(* Logix 5000 project; controller _GigaDiscovery vendor 1 type 14 code 244 rev 35.11; software revision 35.03; part 6 of 23 *)
(* tags used below, declared in another part *)
   Encoder_Pulses : DINT;
   Pignone : DINT;
   Pylon_Axe_Position_360_SUB : REAL;
   Ralla : DINT;
   RallaPignone : REAL;
   Riduttore : REAL;
   Timer : TIMER[50];
   Clock : DINT;   // Base tempi 10 milli sec
   Clock_1_Hz : BOOL;   // SL Clock 1 Hz 0.5 sec OFF 0.5 sec ON
   Clock_4_Hz : BOOL;   // SL Clock 4 Hz 0.125 sec OFF 0.125 sec ON
   Emergency_Brake_manual_Perm : BOOL;
   Emergency_Brake_SL : ALIAS FOR K300_OCC:6:O.6;   // _S31207D
   Gates_Open_Permissive : Permissive;
   Gondola_Axe : Axe;
   HMI_Lamp_Test : BOOL;
   HMI_Monitor_Bars_Time : DINT;
   I_EStop_Pb_OCC1 : UDT_DCI_STOP_TEST;   // +OCC E-stop -S30301F
   I_EStop_Pb_OCC2 : UDT_DCI_STOP_TEST;   // +OCC2 E-Stop -S28502F
   I_Gate_2_Opened : BOOL;   // Gate 2 RFID Sensor Closed -B24601J
   I_Gate_3_Opened : BOOL;   // Gate 3 RFID Sensor Closed -B24701J
   I_Gate_ENTER_G01_Closed : UDT_DCM;   // GATE ENTER (G01) -B25204I
   I_Gate_EXIT_G05_Closed : UDT_DCM;   // GATE EXIT (G05) -B25304I
   I_OCC1_Stop_Cycle_PB : BOOL;   // Stop Cycle -S30308F
   I_OCC2_ACONFIRM : BOOL;   // OCC2 Allow Main CONFIRM -S28602F
   I_OCC2_Stop_Cycle_PB : BOOL;   // Stop Cycle -S28606F
   I_OCC_Emergency_Brake : BOOL;   // I OCC Emergency Brake -S31207D
   I_OCC_Operator_Enable_Key : BOOL;   // OCC Console Enabled -S30305F
   I_Zero_Set_Sensor : BOOL;   // Zero Set Sensor -B11201A
   Impulsi_per_360_gradi : DINT;
   Impulsi_per_grado : REAL;
   K_Speed_Factor : REAL;
   Mem_RESTRAINTS_closed_Correctly : BOOL;
   MODE : BOOL;   // MODE 0 = AUTO 1 = MANUAL -S30801F
   No_Emergencies_CL0 : BOOL;
   No_Emergencies_CL1 : BOOL;
   No_Sfty : Std_to_Sfty;
   O_Close_Gate2 : BOOL;   // Gate 2 Exit Close = Mag ON
   O_Close_Gate3 : BOOL;   // Gate 3 Entrance Close = Mag ON
   O_OCC_EStop_SL : ALIAS FOR K300_OCC:5:O.7;   // -S30301F EMERGENCY
   O_Start_Signal_2 : ALIAS FOR K300_OCC:5:O.2;   // -S30401F RIDE START
   Pb_Platform_Stop : BOOL;   // Platform Stop Command -S30608F
   Platform_Close_Cycle : Sequencer;
   Platform_Close_Permissive_OK : BOOL;
   Platform_Closed_Aux : DINT;
   Platform_Open_Cycle : Sequencer;
   Platform_Open_Permissive : Permissive;
   Platform_Open_Permissive_Ok : BOOL;
   Platform_Opened_Aux : DINT;
   PltaformClosed_CycleComplete : BOOL;   // Piattaforme chiuse e ciclo completato
   PltaformOpeneded_CycleComplete : BOOL;   // Rilevazione Piattaforme aperte con ciclo Completato
   Pylon_Axe : Axe;
   Pylon_Filtered_Speed : REAL;
   Pylon_Filtered_Speed_ABS : REAL;
   Pylon_Stop_Phase : BOOL;
   Reset_Status_SL_Request : BOOL;
   RESTRAINTS_Closed : BOOL;   // All RESTRAINTS Closed
   RESTRAINTS_Open_Postion : BOOL[64];
   RESTRAINTS_Sector : LapBars_Sector[9];
   Start_Platform_AutoCycle_Pylon : BOOL;
   Start_Stop_Cycle : Sequencer;
   Timers : TIMER[32];
   To_Sfty : Std_to_Sfty;
(* Input, continued *)

ROUTINE _04_RESTRAINTS   (* ladder *)
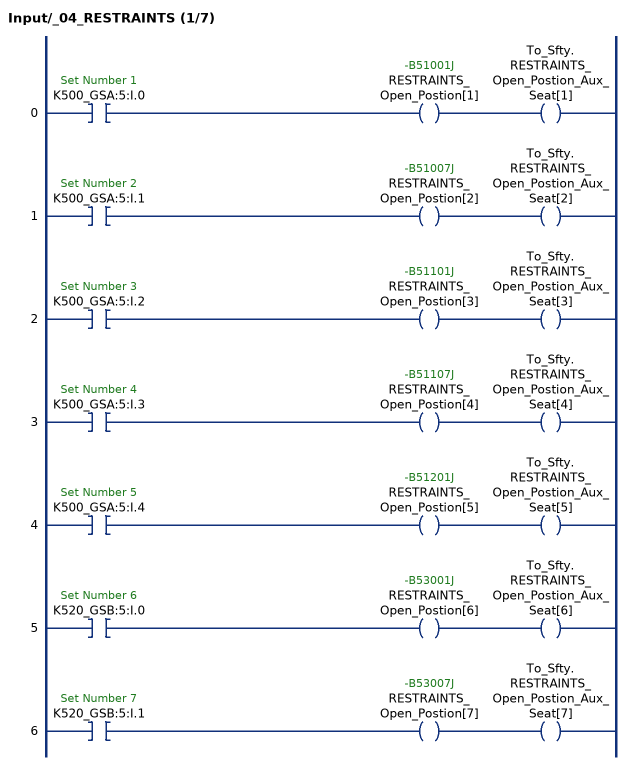
   0: XIC(K500_GSA:5:I.0)OTE(RESTRAINTS_Open_Postion[1])OTE(To_Sfty.RESTRAINTS_Open_Postion_Aux_Seat[1]);
   1: XIC(K500_GSA:5:I.1)OTE(RESTRAINTS_Open_Postion[2])OTE(To_Sfty.RESTRAINTS_Open_Postion_Aux_Seat[2]);
   2: XIC(K500_GSA:5:I.2)OTE(RESTRAINTS_Open_Postion[3])OTE(To_Sfty.RESTRAINTS_Open_Postion_Aux_Seat[3]);
   3: XIC(K500_GSA:5:I.3)OTE(RESTRAINTS_Open_Postion[4])OTE(To_Sfty.RESTRAINTS_Open_Postion_Aux_Seat[4]);
   4: XIC(K500_GSA:5:I.4)OTE(RESTRAINTS_Open_Postion[5])OTE(To_Sfty.RESTRAINTS_Open_Postion_Aux_Seat[5]);
   5: XIC(K520_GSB:5:I.0)OTE(RESTRAINTS_Open_Postion[6])OTE(To_Sfty.RESTRAINTS_Open_Postion_Aux_Seat[6]);
   6: XIC(K520_GSB:5:I.1)OTE(RESTRAINTS_Open_Postion[7])OTE(To_Sfty.RESTRAINTS_Open_Postion_Aux_Seat[7]);
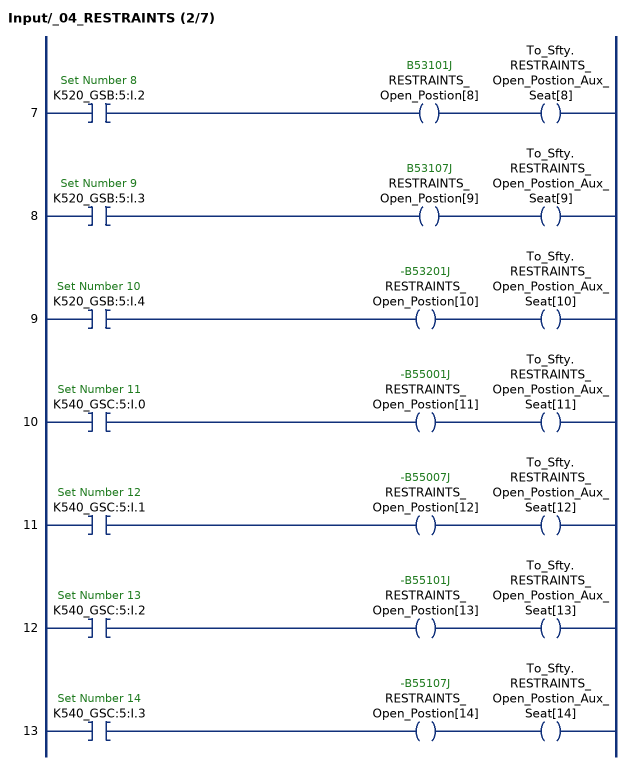
   7: XIC(K520_GSB:5:I.2)OTE(RESTRAINTS_Open_Postion[8])OTE(To_Sfty.RESTRAINTS_Open_Postion_Aux_Seat[8]);
   8: XIC(K520_GSB:5:I.3)OTE(RESTRAINTS_Open_Postion[9])OTE(To_Sfty.RESTRAINTS_Open_Postion_Aux_Seat[9]);
   9: XIC(K520_GSB:5:I.4)OTE(RESTRAINTS_Open_Postion[10])OTE(To_Sfty.RESTRAINTS_Open_Postion_Aux_Seat[10]);
   10: XIC(K540_GSC:5:I.0)OTE(RESTRAINTS_Open_Postion[11])OTE(To_Sfty.RESTRAINTS_Open_Postion_Aux_Seat[11]);
   11: XIC(K540_GSC:5:I.1)OTE(RESTRAINTS_Open_Postion[12])OTE(To_Sfty.RESTRAINTS_Open_Postion_Aux_Seat[12]);
   12: XIC(K540_GSC:5:I.2)OTE(RESTRAINTS_Open_Postion[13])OTE(To_Sfty.RESTRAINTS_Open_Postion_Aux_Seat[13]);
   13: XIC(K540_GSC:5:I.3)OTE(RESTRAINTS_Open_Postion[14])OTE(To_Sfty.RESTRAINTS_Open_Postion_Aux_Seat[14]);
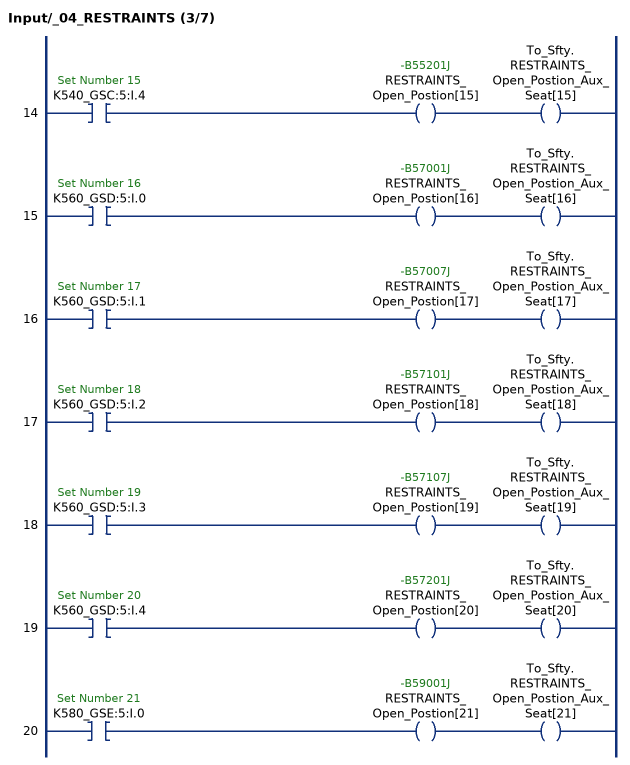
   14: XIC(K540_GSC:5:I.4)OTE(RESTRAINTS_Open_Postion[15])OTE(To_Sfty.RESTRAINTS_Open_Postion_Aux_Seat[15]);
   15: XIC(K560_GSD:5:I.0)OTE(RESTRAINTS_Open_Postion[16])OTE(To_Sfty.RESTRAINTS_Open_Postion_Aux_Seat[16]);
   16: XIC(K560_GSD:5:I.1)OTE(RESTRAINTS_Open_Postion[17])OTE(To_Sfty.RESTRAINTS_Open_Postion_Aux_Seat[17]);
   17: XIC(K560_GSD:5:I.2)OTE(RESTRAINTS_Open_Postion[18])OTE(To_Sfty.RESTRAINTS_Open_Postion_Aux_Seat[18]);
   18: XIC(K560_GSD:5:I.3)OTE(RESTRAINTS_Open_Postion[19])OTE(To_Sfty.RESTRAINTS_Open_Postion_Aux_Seat[19]);
   19: XIC(K560_GSD:5:I.4)OTE(RESTRAINTS_Open_Postion[20])OTE(To_Sfty.RESTRAINTS_Open_Postion_Aux_Seat[20]);
   20: XIC(K580_GSE:5:I.0)OTE(RESTRAINTS_Open_Postion[21])OTE(To_Sfty.RESTRAINTS_Open_Postion_Aux_Seat[21]);
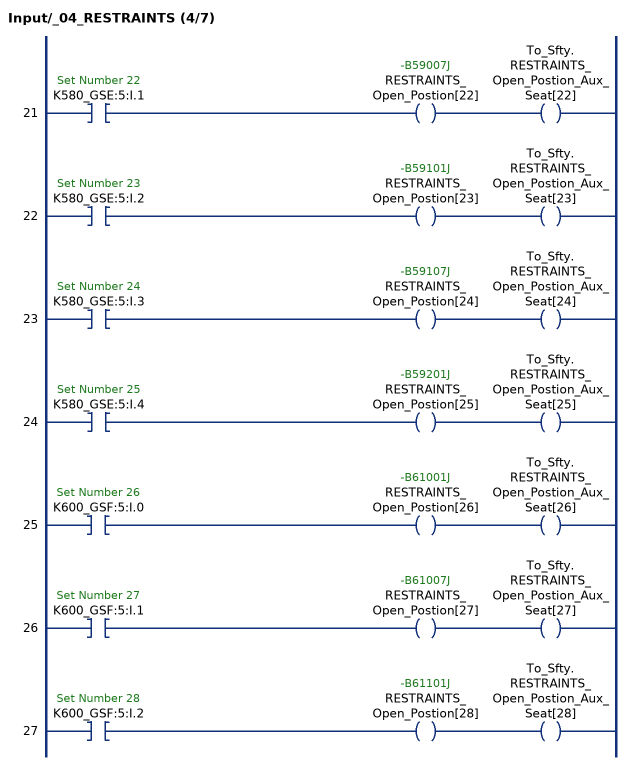
   21: XIC(K580_GSE:5:I.1)OTE(RESTRAINTS_Open_Postion[22])OTE(To_Sfty.RESTRAINTS_Open_Postion_Aux_Seat[22]);
   22: XIC(K580_GSE:5:I.2)OTE(RESTRAINTS_Open_Postion[23])OTE(To_Sfty.RESTRAINTS_Open_Postion_Aux_Seat[23]);
   23: XIC(K580_GSE:5:I.3)OTE(RESTRAINTS_Open_Postion[24])OTE(To_Sfty.RESTRAINTS_Open_Postion_Aux_Seat[24]);
   24: XIC(K580_GSE:5:I.4)OTE(RESTRAINTS_Open_Postion[25])OTE(To_Sfty.RESTRAINTS_Open_Postion_Aux_Seat[25]);
   25: XIC(K600_GSF:5:I.0)OTE(RESTRAINTS_Open_Postion[26])OTE(To_Sfty.RESTRAINTS_Open_Postion_Aux_Seat[26]);
   26: XIC(K600_GSF:5:I.1)OTE(RESTRAINTS_Open_Postion[27])OTE(To_Sfty.RESTRAINTS_Open_Postion_Aux_Seat[27]);
   27: XIC(K600_GSF:5:I.2)OTE(RESTRAINTS_Open_Postion[28])OTE(To_Sfty.RESTRAINTS_Open_Postion_Aux_Seat[28]);
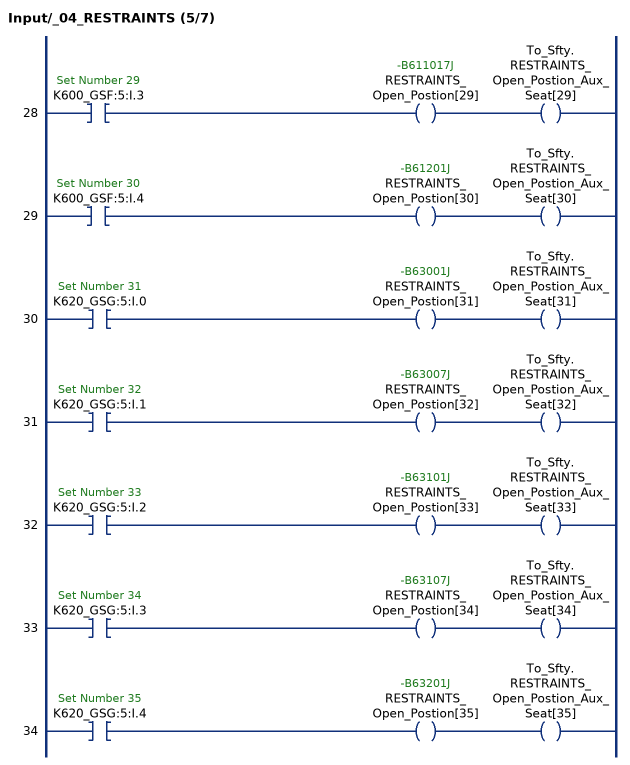
   28: XIC(K600_GSF:5:I.3)OTE(RESTRAINTS_Open_Postion[29])OTE(To_Sfty.RESTRAINTS_Open_Postion_Aux_Seat[29]);
   29: XIC(K600_GSF:5:I.4)OTE(RESTRAINTS_Open_Postion[30])OTE(To_Sfty.RESTRAINTS_Open_Postion_Aux_Seat[30]);
   30: XIC(K620_GSG:5:I.0)OTE(RESTRAINTS_Open_Postion[31])OTE(To_Sfty.RESTRAINTS_Open_Postion_Aux_Seat[31]);
   31: XIC(K620_GSG:5:I.1)OTE(RESTRAINTS_Open_Postion[32])OTE(To_Sfty.RESTRAINTS_Open_Postion_Aux_Seat[32]);
   32: XIC(K620_GSG:5:I.2)OTE(RESTRAINTS_Open_Postion[33])OTE(To_Sfty.RESTRAINTS_Open_Postion_Aux_Seat[33]);
   33: XIC(K620_GSG:5:I.3)OTE(RESTRAINTS_Open_Postion[34])OTE(To_Sfty.RESTRAINTS_Open_Postion_Aux_Seat[34]);
   34: XIC(K620_GSG:5:I.4)OTE(RESTRAINTS_Open_Postion[35])OTE(To_Sfty.RESTRAINTS_Open_Postion_Aux_Seat[35]);
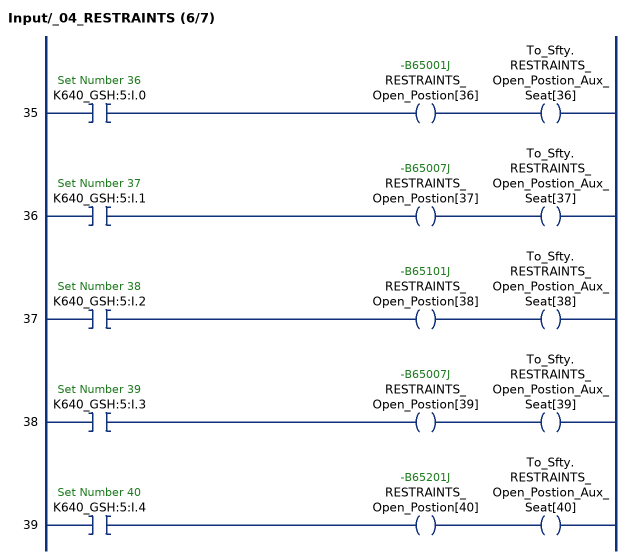
   35: XIC(K640_GSH:5:I.0)OTE(RESTRAINTS_Open_Postion[36])OTE(To_Sfty.RESTRAINTS_Open_Postion_Aux_Seat[36]);
   36: XIC(K640_GSH:5:I.1)OTE(RESTRAINTS_Open_Postion[37])OTE(To_Sfty.RESTRAINTS_Open_Postion_Aux_Seat[37]);
   37: XIC(K640_GSH:5:I.2)OTE(RESTRAINTS_Open_Postion[38])OTE(To_Sfty.RESTRAINTS_Open_Postion_Aux_Seat[38]);
   38: XIC(K640_GSH:5:I.3)OTE(RESTRAINTS_Open_Postion[39])OTE(To_Sfty.RESTRAINTS_Open_Postion_Aux_Seat[39]);
   39: XIC(K640_GSH:5:I.4)OTE(RESTRAINTS_Open_Postion[40])OTE(To_Sfty.RESTRAINTS_Open_Postion_Aux_Seat[40]);
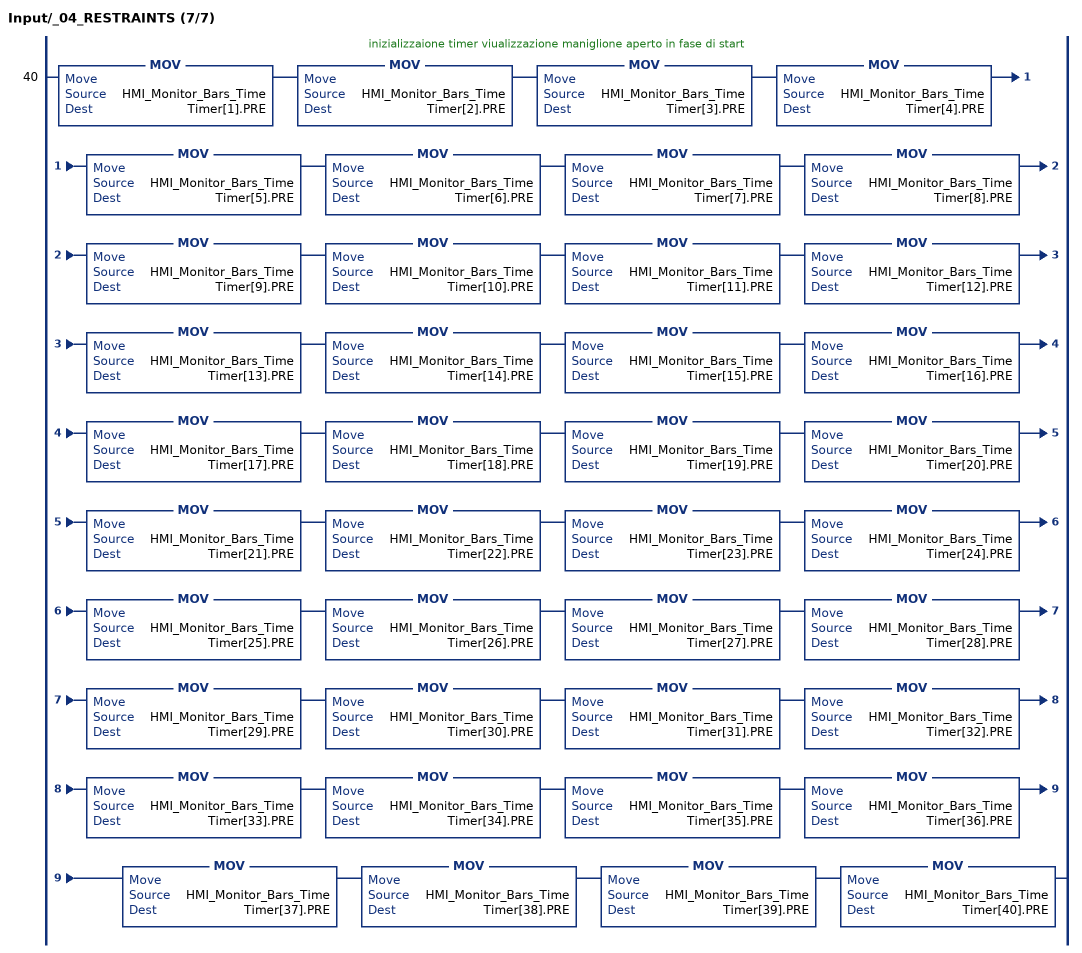
   // inizializzaione timer viualizzazione maniglione aperto in fase di start
   40: MOV(HMI_Monitor_Bars_Time,Timer[1].PRE)MOV(HMI_Monitor_Bars_Time,Timer[2].PRE)MOV(HMI_Monitor_Bars_Time,Timer[3].PRE)MOV(HMI_Monitor_Bars_Time,Timer[4].PRE)MOV(HMI_Monitor_Bars_Time,Timer[5].PRE)MOV(HMI_Monitor_Bars_Time,Timer[6].PRE)MOV(HMI_Monitor_Bars_Time,Timer[7].PRE)MOV(HMI_Monitor_Bars_Time,Timer[8].PRE)MOV(HMI_Monitor_Bars_Time,Timer[9].PRE)MOV(HMI_Monitor_Bars_Time,Timer[10].PRE)MOV(HMI_Monitor_Bars_Time,Timer[11].PRE)MOV(HMI_Monitor_Bars_Time,Timer[12].PRE)MOV(HMI_Monitor_Bars_Time,Timer[13].PRE)MOV(HMI_Monitor_Bars_Time,Timer[14].PRE)MOV(HMI_Monitor_Bars_Time,Timer[15].PRE)MOV(HMI_Monitor_Bars_Time,Timer[16].PRE)MOV(HMI_Monitor_Bars_Time,Timer[17].PRE)MOV(HMI_Monitor_Bars_Time,Timer[18].PRE)MOV(HMI_Monitor_Bars_Time,Timer[19].PRE)MOV(HMI_Monitor_Bars_Time,Timer[20].PRE)MOV(HMI_Monitor_Bars_Time,Timer[21].PRE)MOV(HMI_Monitor_Bars_Time,Timer[22].PRE)MOV(HMI_Monitor_Bars_Time,Timer[23].PRE)MOV(HMI_Monitor_Bars_Time,Timer[24].PRE)MOV(HMI_Monitor_Bars_Time,Timer[25].PRE)MOV(HMI_Monitor_Bars_Time,Timer[26].PRE)MOV(HMI_Monitor_Bars_Time,Timer[27].PRE)MOV(HMI_Monitor_Bars_Time,Timer[28].PRE)MOV(HMI_Monitor_Bars_Time,Timer[29].PRE)MOV(HMI_Monitor_Bars_Time,Timer[30].PRE)MOV(HMI_Monitor_Bars_Time,Timer[31].PRE)MOV(HMI_Monitor_Bars_Time,Timer[32].PRE)MOV(HMI_Monitor_Bars_Time,Timer[33].PRE)MOV(HMI_Monitor_Bars_Time,Timer[34].PRE)MOV(HMI_Monitor_Bars_Time,Timer[35].PRE)MOV(HMI_Monitor_Bars_Time,Timer[36].PRE)MOV(HMI_Monitor_Bars_Time,Timer[37].PRE)MOV(HMI_Monitor_Bars_Time,Timer[38].PRE)MOV(HMI_Monitor_Bars_Time,Timer[39].PRE)MOV(HMI_Monitor_Bars_Time,Timer[40].PRE);
END_ROUTINE

ROUTINE _05_Platform   (* ladder *)
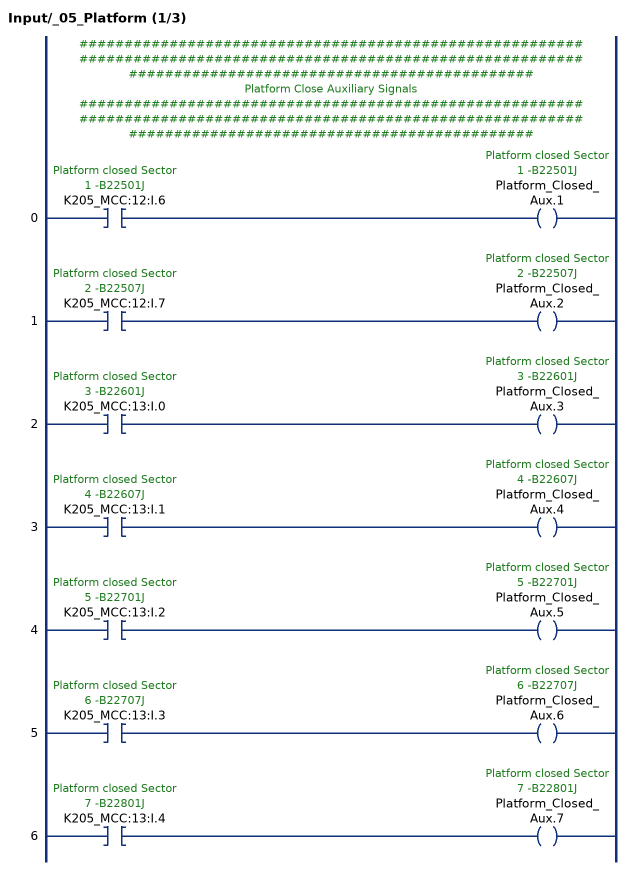
   // #############################################################################################################################################################
   // Platform Close Auxiliary Signals
   // #############################################################################################################################################################
   0: XIC(K205_MCC:12:I.6)OTE(Platform_Closed_Aux.1);
   1: XIC(K205_MCC:12:I.7)OTE(Platform_Closed_Aux.2);
   2: XIC(K205_MCC:13:I.0)OTE(Platform_Closed_Aux.3);
   3: XIC(K205_MCC:13:I.1)OTE(Platform_Closed_Aux.4);
   4: XIC(K205_MCC:13:I.2)OTE(Platform_Closed_Aux.5);
   5: XIC(K205_MCC:13:I.3)OTE(Platform_Closed_Aux.6);
   6: XIC(K205_MCC:13:I.4)OTE(Platform_Closed_Aux.7);
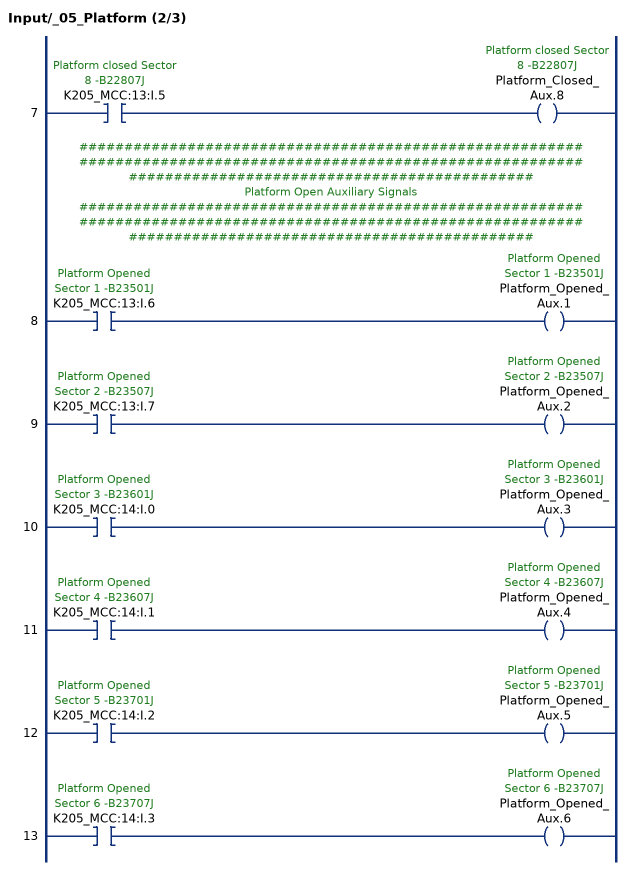
   7: XIC(K205_MCC:13:I.5)OTE(Platform_Closed_Aux.8);
   // #############################################################################################################################################################
   // Platform Open Auxiliary Signals
   // #############################################################################################################################################################
   8: XIC(K205_MCC:13:I.6)OTE(Platform_Opened_Aux.1);
   9: XIC(K205_MCC:13:I.7)OTE(Platform_Opened_Aux.2);
   10: XIC(K205_MCC:14:I.0)OTE(Platform_Opened_Aux.3);
   11: XIC(K205_MCC:14:I.1)OTE(Platform_Opened_Aux.4);
   12: XIC(K205_MCC:14:I.2)OTE(Platform_Opened_Aux.5);
   13: XIC(K205_MCC:14:I.3)OTE(Platform_Opened_Aux.6);
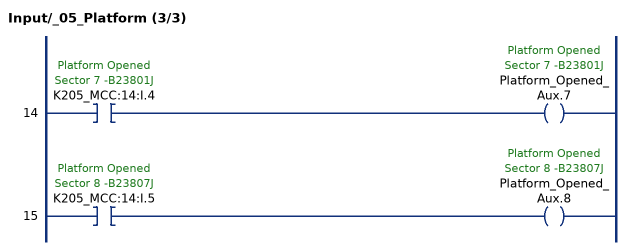
   14: XIC(K205_MCC:14:I.4)OTE(Platform_Opened_Aux.7);
   15: XIC(K205_MCC:14:I.5)OTE(Platform_Opened_Aux.8);
END_ROUTINE

ROUTINE _06_Pylon   (* ladder *)
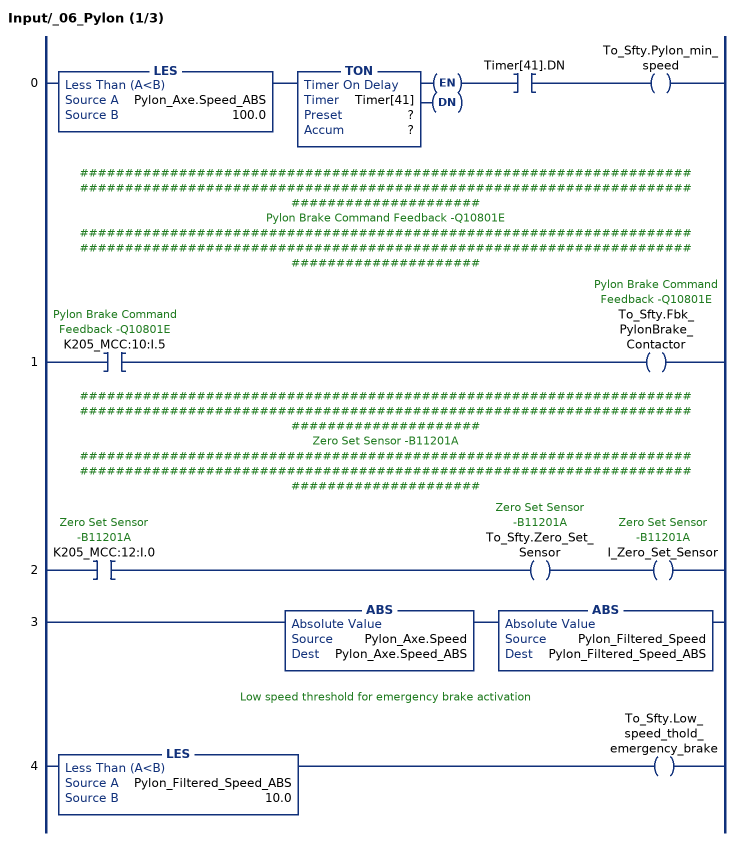
   0: LES(Pylon_Axe.Speed_ABS,100.0)TON(Timer[41],?,?)XIC(Timer[41].DN)OTE(To_Sfty.Pylon_min_speed);
   // #############################################################################################################################################################
   // Pylon Brake Command Feedback -Q10801E
   // #############################################################################################################################################################
   1: XIC(K205_MCC:10:I.5)OTE(To_Sfty.Fbk_PylonBrake_Contactor);
   // #############################################################################################################################################################
   // Zero Set Sensor -B11201A
   // #############################################################################################################################################################
   2: XIC(K205_MCC:12:I.0)OTE(To_Sfty.Zero_Set_Sensor)OTE(I_Zero_Set_Sensor);
   3: ABS(Pylon_Axe.Speed,Pylon_Axe.Speed_ABS)ABS(Pylon_Filtered_Speed,Pylon_Filtered_Speed_ABS);
   // Low speed threshold for emergency brake activation
   4: LES(Pylon_Filtered_Speed_ABS,10.0)OTE(To_Sfty.Low_speed_thold_emergency_brake);
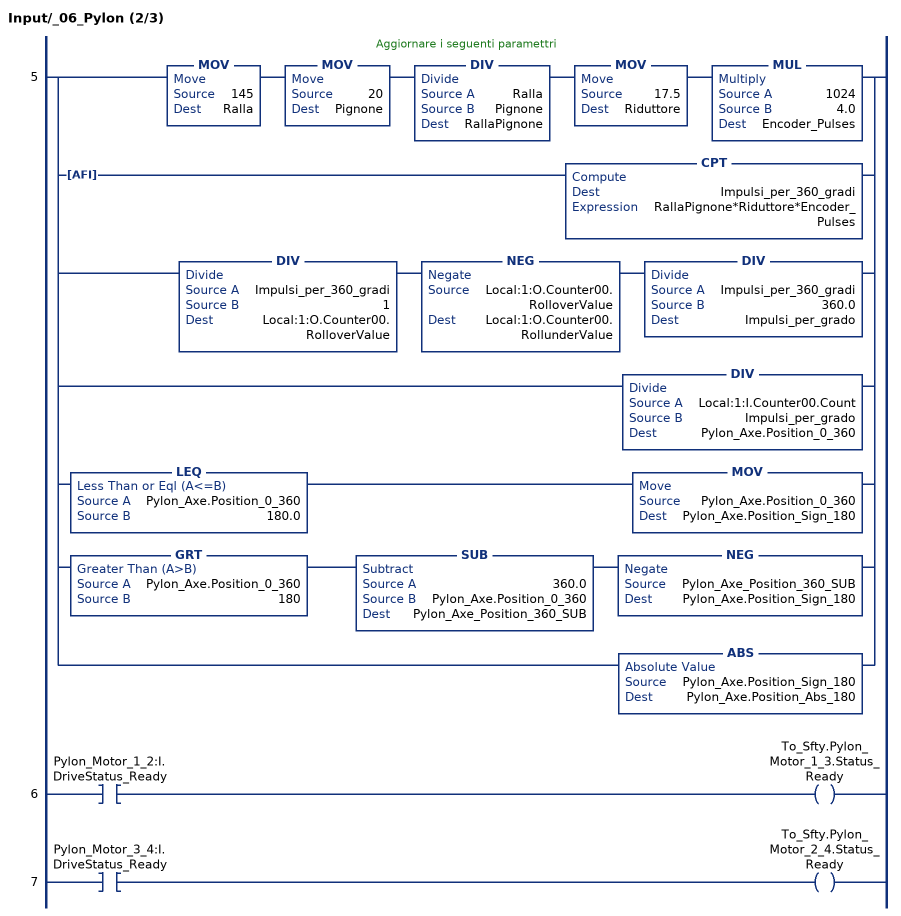
   // Aggiornare i seguenti paramettri
   5: [MOV(145,Ralla) MOV(20,Pignone) DIV(Ralla,Pignone,RallaPignone) MOV(17.5,Riduttore) MUL(1024,4.0,Encoder_Pulses) ,AFI() CPT(Impulsi_per_360_gradi,RallaPignone*Riduttore*Encoder_Pulses) ,DIV(Impulsi_per_360_gradi,1,Local:1:O.Counter00.RolloverValue) NEG(Local:1:O.Counter00.RolloverValue,Local:1:O.Counter00.RollunderValue) DIV(Impulsi_per_360_gradi,360.0,Impulsi_per_grado) ,DIV(Local:1:I.Counter00.Count,Impulsi_per_grado,Pylon_Axe.Position_0_360) ,LEQ(Pylon_Axe.Position_0_360,180.0) MOV(Pylon_Axe.Position_0_360,Pylon_Axe.Position_Sign_180) ,GRT(Pylon_Axe.Position_0_360,180) SUB(360.0,Pylon_Axe.Position_0_360,Pylon_Axe_Position_360_SUB) NEG(Pylon_Axe_Position_360_SUB,Pylon_Axe.Position_Sign_180) ,ABS(Pylon_Axe.Position_Sign_180,Pylon_Axe.Position_Abs_180) ];
   6: XIC(Pylon_Motor_1_2:I.DriveStatus_Ready)OTE(To_Sfty.Pylon_Motor_1_3.Status_Ready);
   7: XIC(Pylon_Motor_3_4:I.DriveStatus_Ready)OTE(To_Sfty.Pylon_Motor_2_4.Status_Ready);
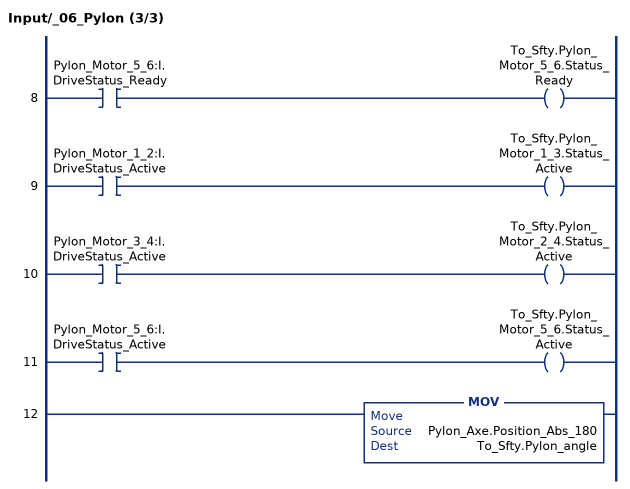
   8: XIC(Pylon_Motor_5_6:I.DriveStatus_Ready)OTE(To_Sfty.Pylon_Motor_5_6.Status_Ready);
   9: XIC(Pylon_Motor_1_2:I.DriveStatus_Active)OTE(To_Sfty.Pylon_Motor_1_3.Status_Active);
   10: XIC(Pylon_Motor_3_4:I.DriveStatus_Active)OTE(To_Sfty.Pylon_Motor_2_4.Status_Active);
   11: XIC(Pylon_Motor_5_6:I.DriveStatus_Active)OTE(To_Sfty.Pylon_Motor_5_6.Status_Active);
   12: MOV(Pylon_Axe.Position_Abs_180,To_Sfty.Pylon_angle);
END_ROUTINE

ROUTINE _07_Gondola   (* ladder *)
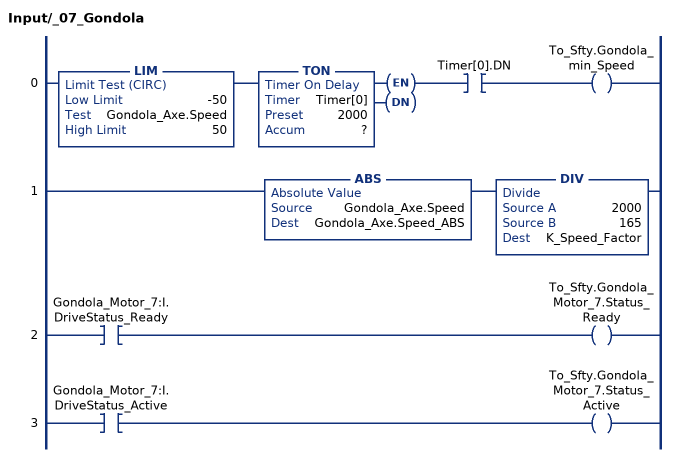
   0: LIM(-50,Gondola_Axe.Speed,50)TON(Timer[0],?,?)XIC(Timer[0].DN)OTE(To_Sfty.Gondola_min_Speed);
   1: ABS(Gondola_Axe.Speed,Gondola_Axe.Speed_ABS)DIV(2000,165,K_Speed_Factor);
   2: XIC(Gondola_Motor_7:I.DriveStatus_Ready)OTE(To_Sfty.Gondola_Motor_7.Status_Ready);
   3: XIC(Gondola_Motor_7:I.DriveStatus_Active)OTE(To_Sfty.Gondola_Motor_7.Status_Active);
END_ROUTINE

ROUTINE Main   (* ladder *)
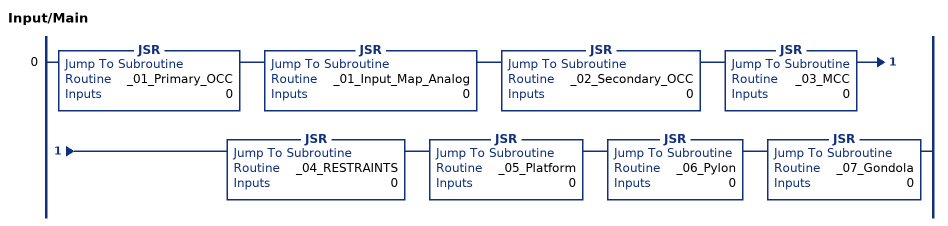
   0: JSR(_01_Primary_OCC,0)JSR(_01_Input_Map_Analog,0)JSR(_02_Secondary_OCC,0)JSR(_03_MCC,0)JSR(_04_RESTRAINTS,0)JSR(_05_Platform,0)JSR(_06_Pylon,0)JSR(_07_Gondola,0);
END_ROUTINE
END_PROGRAM

PROGRAM Main10ms   (* main routine Main *)

ROUTINE Main   (* ladder *)
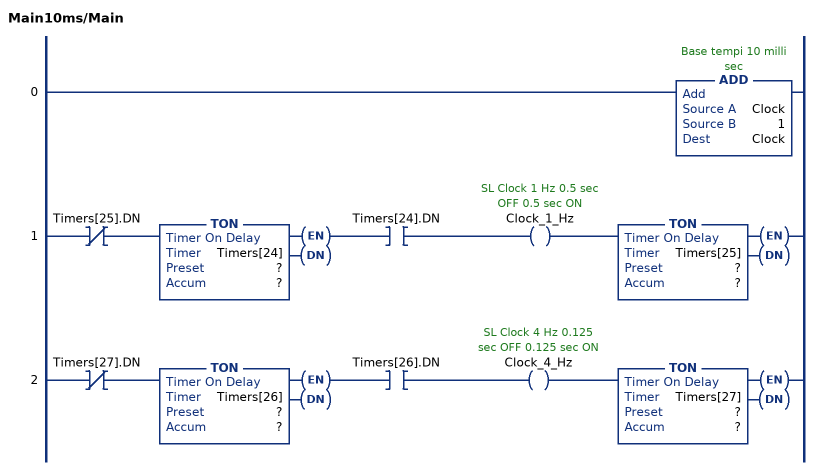
   0: ADD(Clock,1,Clock);
   1: XIO(Timers[25].DN)TON(Timers[24],?,?)XIC(Timers[24].DN)OTE(Clock_1_Hz)TON(Timers[25],?,?);
   2: XIO(Timers[27].DN)TON(Timers[26],?,?)XIC(Timers[26].DN)OTE(Clock_4_Hz)TON(Timers[27],?,?);
END_ROUTINE
END_PROGRAM

PROGRAM Output   (* main routine Main *)
VAR
   EntryGate : Sfq_Lamp := (Input := 1, LampCoil := 1);
   ExitGate : Sfq_Lamp := (Input := 1, LampCoil := 1);
   I_OCC1_Stop_Cycle_PB_memory : BOOL;
   I_OCC2_Stop_Cycle_PB_memory : BOOL;
   O_Alarm_Noise : BOOL;
   O_Alarm_Signal : BOOL;
   O_Allow_Operator : BOOL;
   O_ExitGate_Signal : BOOL := 1;
   O_Lapbars_Open : ALIAS FOR K300_OCC:5:O.4;
   O_Platform_Close_Signal : ALIAS FOR K300_OCC:5:O.6;   // -S30605F PLATFORM CLOSING
   O_Platform_Open_Signal : ALIAS FOR K300_OCC:5:O.5;   // -S30601F PLATFORM OPENING
   O_Start_Signal : ALIAS FOR K300_OCC:5:O.1;   // -S30403F RIDE START
   O_Stop_Signal : ALIAS FOR K300_OCC:5:O.0;   // -S30308F RIDE STOP
   Os : DINT;
   Out_FGEN_01 : FUNCTION_GENERATOR := (XY1Size := 2, Out := -90.0);
   Out_FGEN_06 : FUNCTION_GENERATOR := (XY1Size := 2);
   Out_FGEN_07 : FUNCTION_GENERATOR := (In := -1.0, XY1Size := 2);
   Out_FGEN_09 : FUNCTION_GENERATOR := (XY1Size := 2);
   Out_FGEN_10 : FUNCTION_GENERATOR := (In := 100.0, XY1Size := 2, Out := 10000.0);
   Output_Scalaggi : Scale_2_P[16] := ([0].Input[1] := 100.0, [0].Output[0] := -90.0, [0].Output[1] := 90.0, [1].Input[0] := -100.0, [1].Input[1] := 100.0, [1].Output[0] := -10000.0, [1].Output[1] := 10000.0, [2].Input[1] := 100.0, [2].Output[1] := 10000.0, [3].Input[0] := -100.0, [3].Input[1] := 100.0, [3].Output[0] := -10000.0, [3].Output[1] := 10000.0, [4].Input[1] := 31218.0, [4].Output[1] := 10.0, [5].Input[1] := 31218.0, [5].Output[1] := 10.0, [6].Input[1] := 31218.0, [6].Output[1] := 10.0, [7].Input[1] := 31218.0, [7].Output[1] := 10.0, [8].Input[1] := 31218.0, [8].Output[1] := 10.0, [9].Input[1] := 31218.0, [9].Output[1] := 10.0, [11].Input[0] := -1.0, [11].Input[1] := 1.0, [11].Output[1] := 10000.0, [12].Input[0] := -1.0, [12].Input[1] := 1.0, [12].Output[0] := -10000.0, [12].Output[1] := 10000.0);
   RAD_01 : FBD_MATH_ADVANCED := (Source := -90.0, Dest := -1.5707964);
   SFQ_disable : BOOL;
   SFQ_Mask : DINT := -269484034;
   SFQ_Mask2 : DINT;
   SFQ_MASK_OK : DINT := -1;
   SFQBit : BOOL;
   SIN_01 : FBD_MATH_ADVANCED := (Source := -1.5707964, Dest := -1.0);
   Start_Permissive_MakCompare : DINT := -1048577;
   TempSFQ : DINT;
END_VAR

ROUTINE _01_Primary_OCC   (* ladder *)
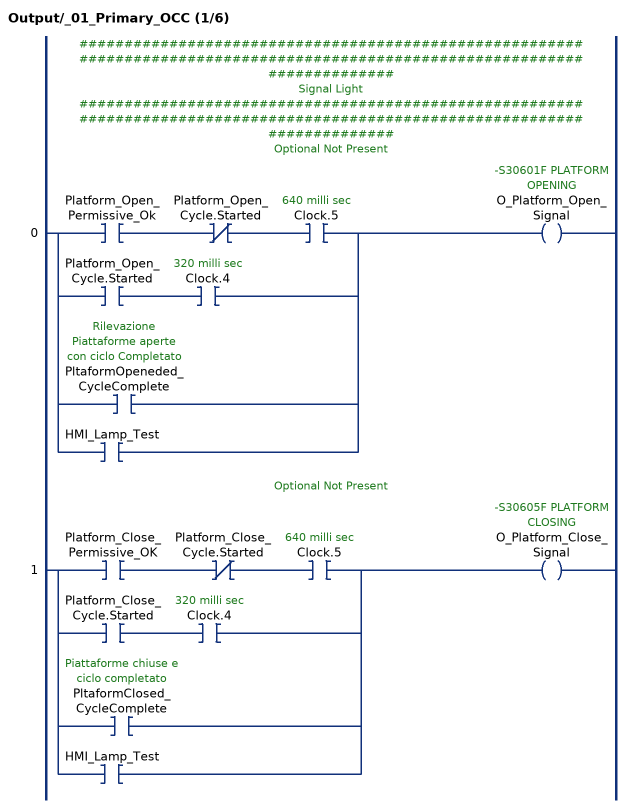
   // ##############################################################################################################################
   // Signal Light
   // ##############################################################################################################################
   // Optional Not Present
   0: [XIC(Platform_Open_Permissive_Ok) XIO(Platform_Open_Cycle.Started) XIC(Clock.5) ,XIC(Platform_Open_Cycle.Started) XIC(Clock.4) ,XIC(PltaformOpeneded_CycleComplete) ,XIC(HMI_Lamp_Test) ]OTE(O_Platform_Open_Signal);
   // Optional Not Present
   1: [XIC(Platform_Close_Permissive_OK) XIO(Platform_Close_Cycle.Started) XIC(Clock.5) ,XIC(Platform_Close_Cycle.Started) XIC(Clock.4) ,XIC(PltaformClosed_CycleComplete) ,XIC(HMI_Lamp_Test) ]OTE(O_Platform_Close_Signal);
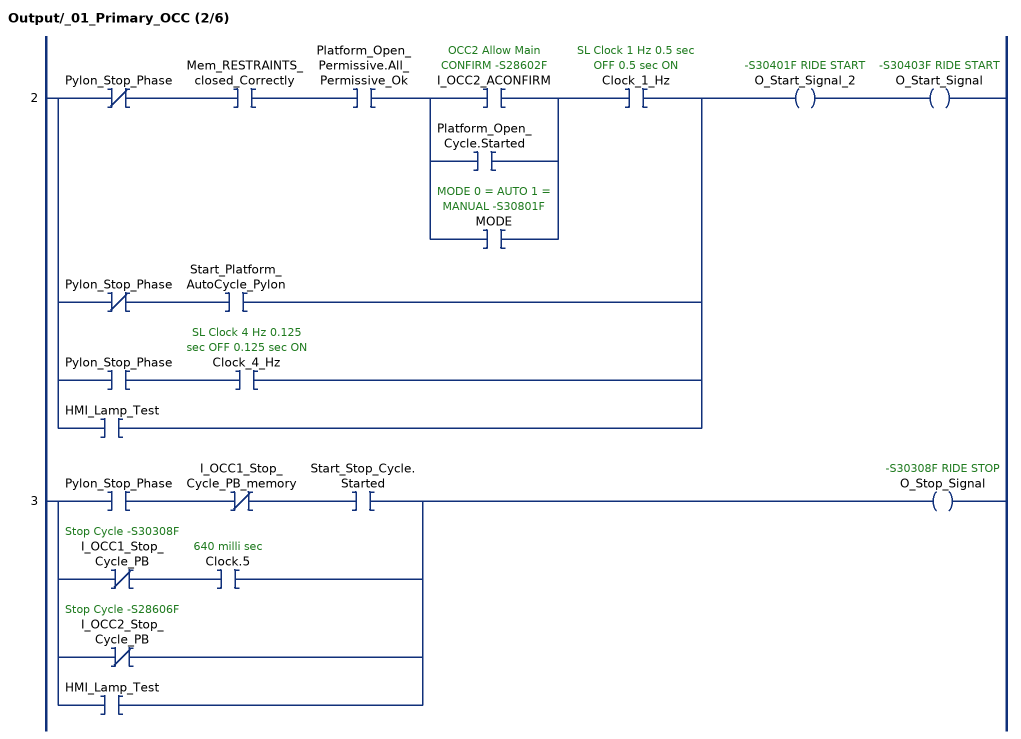
   2: [XIO(Pylon_Stop_Phase) XIC(Mem_RESTRAINTS_closed_Correctly) XIC(Platform_Open_Permissive.All_Permissive_Ok) [XIC(I_OCC2_ACONFIRM) ,XIC(Platform_Open_Cycle.Started) ,XIC(MODE) ] XIC(Clock_1_Hz) ,XIO(Pylon_Stop_Phase) XIC(Start_Platform_AutoCycle_Pylon) ,XIC(Pylon_Stop_Phase) XIC(Clock_4_Hz) ,XIC(HMI_Lamp_Test) ]OTE(O_Start_Signal_2)OTE(O_Start_Signal);
   3: [XIC(Pylon_Stop_Phase) XIO(I_OCC1_Stop_Cycle_PB_memory) XIC(Start_Stop_Cycle.Started) ,XIO(I_OCC1_Stop_Cycle_PB) XIC(Clock.5) ,XIO(I_OCC2_Stop_Cycle_PB) ,XIC(HMI_Lamp_Test) ]OTE(O_Stop_Signal);
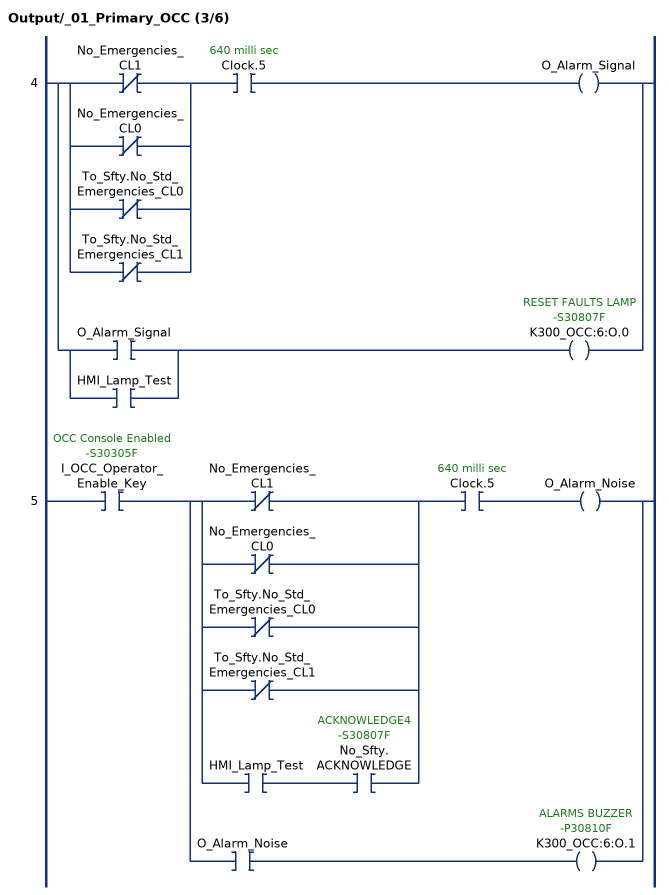
   4: [[XIO(No_Emergencies_CL1) ,XIO(No_Emergencies_CL0) ,XIO(To_Sfty.No_Std_Emergencies_CL0) ,XIO(To_Sfty.No_Std_Emergencies_CL1) ] XIC(Clock.5) OTE(O_Alarm_Signal) ,[XIC(O_Alarm_Signal) ,XIC(HMI_Lamp_Test) ] OTE(K300_OCC:6:O.0) ];
   5: XIC(I_OCC_Operator_Enable_Key)[[XIO(No_Emergencies_CL1) ,XIO(No_Emergencies_CL0) ,XIO(To_Sfty.No_Std_Emergencies_CL0) ,XIO(To_Sfty.No_Std_Emergencies_CL1) ,XIC(HMI_Lamp_Test) XIC(No_Sfty.ACKNOWLEDGE) ] XIC(Clock.5) OTE(O_Alarm_Noise) ,XIC(O_Alarm_Noise) OTE(K300_OCC:6:O.1) ];
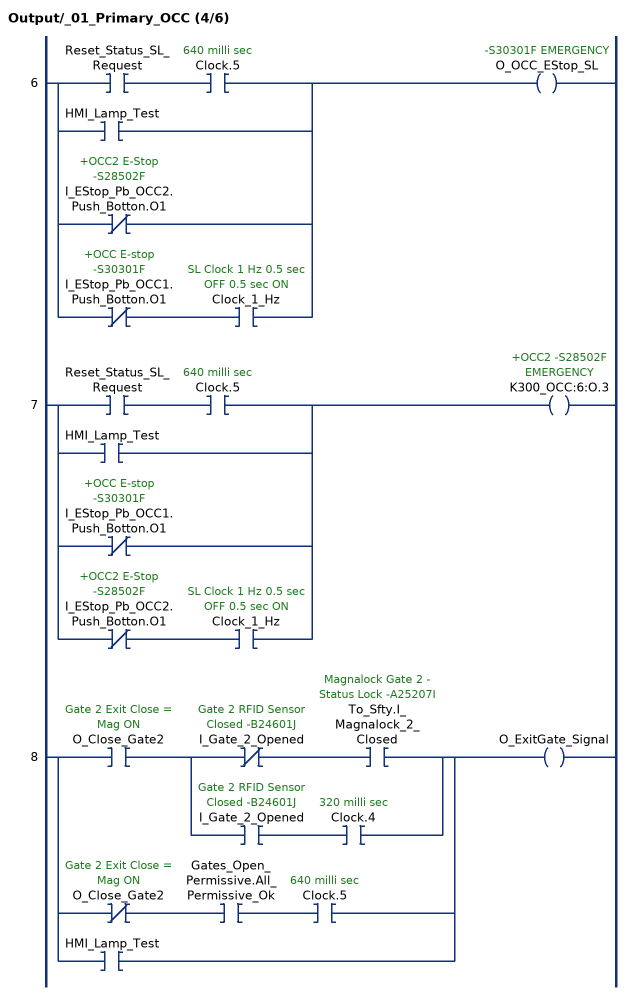
   6: [[XIC(Reset_Status_SL_Request) XIC(Clock.5) ,XIC(HMI_Lamp_Test) ] ,XIO(I_EStop_Pb_OCC2.Push_Botton.O1) ,XIO(I_EStop_Pb_OCC1.Push_Botton.O1) XIC(Clock_1_Hz) ]OTE(O_OCC_EStop_SL);
   7: [[XIC(Reset_Status_SL_Request) XIC(Clock.5) ,XIC(HMI_Lamp_Test) ] ,XIO(I_EStop_Pb_OCC1.Push_Botton.O1) ,XIO(I_EStop_Pb_OCC2.Push_Botton.O1) XIC(Clock_1_Hz) ]OTE(K300_OCC:6:O.3);
   8: [XIC(O_Close_Gate2) [XIO(I_Gate_2_Opened) XIC(To_Sfty.I_Magnalock_2_Closed) ,XIC(I_Gate_2_Opened) XIC(Clock.4) ] ,XIO(O_Close_Gate2) XIC(Gates_Open_Permissive.All_Permissive_Ok) XIC(Clock.5) ,XIC(HMI_Lamp_Test) ]OTE(O_ExitGate_Signal);
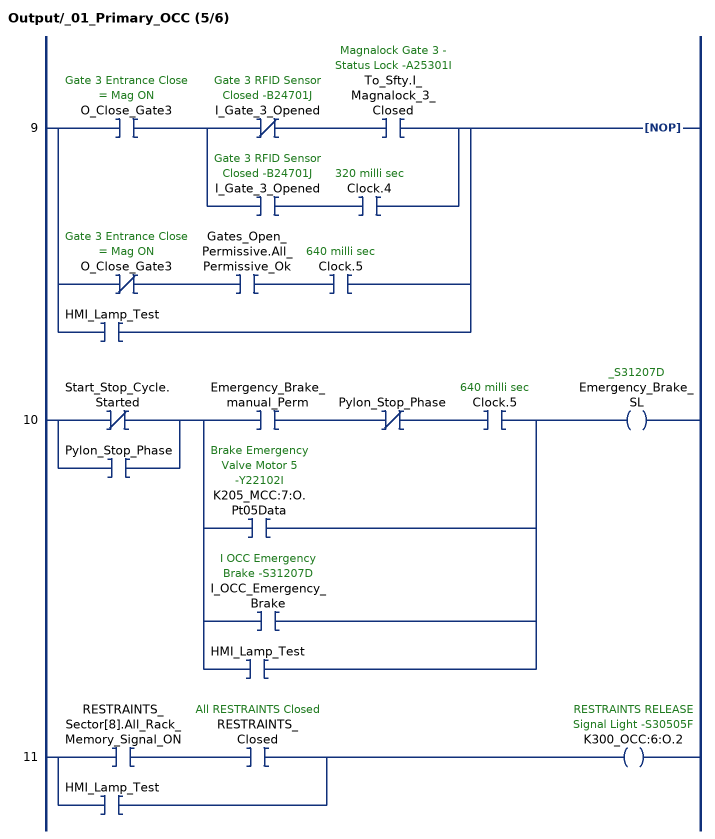
   9: [XIC(O_Close_Gate3) [XIO(I_Gate_3_Opened) XIC(To_Sfty.I_Magnalock_3_Closed) ,XIC(I_Gate_3_Opened) XIC(Clock.4) ] ,XIO(O_Close_Gate3) XIC(Gates_Open_Permissive.All_Permissive_Ok) XIC(Clock.5) ,XIC(HMI_Lamp_Test) ]NOP();
   10: [XIO(Start_Stop_Cycle.Started) ,XIC(Pylon_Stop_Phase) ][XIC(Emergency_Brake_manual_Perm) XIO(Pylon_Stop_Phase) XIC(Clock.5) ,XIC(K205_MCC:7:O.Pt05Data) ,XIC(I_OCC_Emergency_Brake) ,XIC(HMI_Lamp_Test) ]OTE(Emergency_Brake_SL);
   11: [XIC(RESTRAINTS_Sector[8].All_Rack_Memory_Signal_ON) XIC(RESTRAINTS_Closed) ,XIC(HMI_Lamp_Test) ]OTE(K300_OCC:6:O.2);
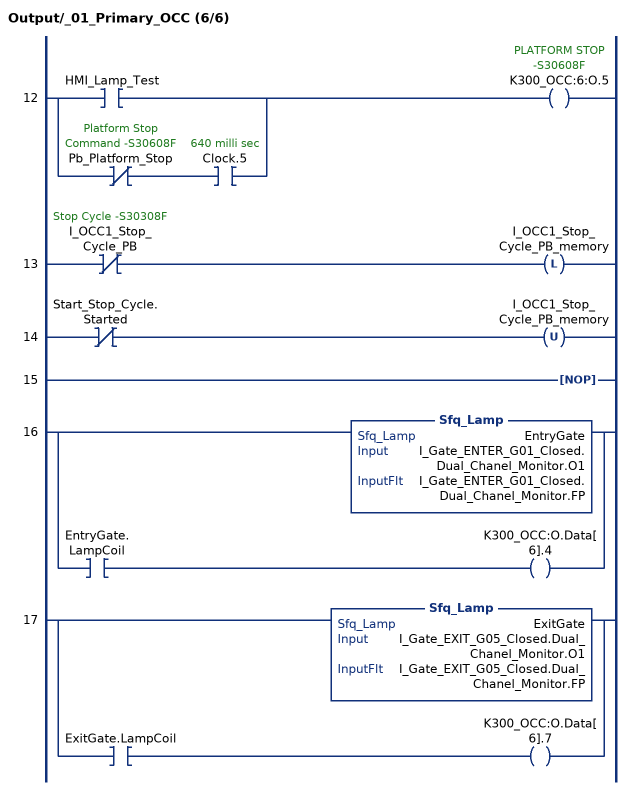
   12: [XIC(HMI_Lamp_Test) ,XIO(Pb_Platform_Stop) XIC(Clock.5) ]OTE(K300_OCC:6:O.5);
   13: XIO(I_OCC1_Stop_Cycle_PB)OTL(I_OCC1_Stop_Cycle_PB_memory);
   14: XIO(Start_Stop_Cycle.Started)OTU(I_OCC1_Stop_Cycle_PB_memory);
   15: NOP();
   16: [Sfq_Lamp(EntryGate,I_Gate_ENTER_G01_Closed.Dual_Chanel_Monitor.O1,I_Gate_ENTER_G01_Closed.Dual_Chanel_Monitor.FP) ,XIC(EntryGate.LampCoil) OTE(K300_OCC:O.Data[6].4) ];
   17: [Sfq_Lamp(ExitGate,I_Gate_EXIT_G05_Closed.Dual_Chanel_Monitor.O1,I_Gate_EXIT_G05_Closed.Dual_Chanel_Monitor.FP) ,XIC(ExitGate.LampCoil) OTE(K300_OCC:O.Data[6].7) ];
END_ROUTINE
